(* Logix 5000 project; controller _GigaDiscovery vendor 1 type 14 code 244 rev 35.11; software revision 35.03; part 4 of 23 *)
(* tags used below, declared in another part *)
   Clock : DINT;   // Base tempi 10 milli sec
   Current_TimeInStation : DINT;
   Cycle_End_Timer : TIMER;
   Cycle_Timing : TIMER;
   Gates_Open_Permissive : Permissive;
   HMI_Angle : REAL;
   HMI_button_addtoindex : BOOL;
   HMI_button_subtracttoindex : BOOL;
   HMI_Current_Screen : DINT;
   HMI_Disable_external_acces : BOOL;   // ROUTER A72A07D Disable external acces
   HMI_Enable_external_acces : BOOL;   // ROUTER A72A07D Eneble external acces
   HMI_JM_Stats_Hist : Run_Count_Hist_JM[10];
   HMI_Lamp_Test : BOOL;
   HMI_Remote_Display : DINT;   // Display control 0 = operator 0 <> PLC
   HMI_Remote_Status : DINT;   // 0 = Disabled 1 = Enable but not remote control 2 = Remote control active
   HMI_Update_Time : BOOL;
   I_Light_Selector : BOOL;   // Light Selector Switch -S30408F
   I_OCC_Operator_Enable_Key : BOOL;   // OCC Console Enabled -S30305F
   I_Remote_Connection_Enabled : BOOL;   // Remote Connection active ROUTER eWON K74A04E
   index_for_stats_hist : DINT;
   Life_of_Machine : Life_of_Machine;
   No_Sfty : Std_to_Sfty;
   O_Enable_Remote_Connection : BOOL;   // ROUTER A72A07D Eneble external acces
   O_Front_Leg_Light : BOOL;   // Fron leg and front light signal -K3204H
   O_Gondola_Pendolum_Light : BOOL;   // Gondola and pendulum light signal -K3206H
   O_Rear_Leg_Light : BOOL;   // Rear leg and rear light signal -K3202H
   Platform_Close_Cycle : Sequencer;
   Platform_Close_Permissive : Permissive;
   Platform_Open_Cycle : Sequencer;
   Platform_Open_Permissive : Permissive;
   PltaformClosed_CycleComplete : BOOL;   // Piattaforme chiuse e ciclo completato
   PltaformOpeneded_CycleComplete : BOOL;   // Rilevazione Piattaforme aperte con ciclo Completato
   Previous_TimeInStation : DINT;
   ProofTest_Req : BOOL;
   RESTRAINTS_Closed : BOOL;   // All RESTRAINTS Closed
   RESTRAINTS_Closing : BOOL;
   Restraints_Cycle : Sequencer;
   RESTRAINTS_Opening : BOOL;
   Restraints_Permissive : Permissive;
   Restraints_Permissive_Ok : BOOL;
   Start_Permissive : Permissive;
   Start_Stop_Cycle : Sequencer;
   Start_TOF : TIMER;
   Stats_Times : DINT[30];
   TimeInStation_Count_Daily : COUNTER;
   TimeInStation_Count_Hourly : COUNTER;
   TimeInStation_Timer : TIMER;   // 10 min 600 sec
   Timers : TIMER[32];
   To_Sfty : Std_to_Sfty;

        [68].time_avg[17] := 29, [68].time_avg[18] := 26, [69].date[0] := -2, [69].date[1] := 1, [69].date[2] := 11, [69].runs[0] := 114, [69].runs[7] := 7, [69].runs[9] := 2, [69].runs[10] := 8, [69].runs[11] := 3, [69].runs[13] := 6, [69].runs[14] := 11, [69].time_avg[0] := 84, [69].time_avg[2] := 22683, [69].time_avg[4] := 28480, [69].time_avg[5] := 22361, [69].time_avg[7] := 107, [69].time_avg[11] := 24, [69].time_avg[13] := 70, [69].time_avg[14] := 104, [70].date[0] := -2, [70].date[1] := 1, [70].date[2] := 8, [70].runs[0] := 19, [70].runs[23] := 3, [70].time_avg[0] := 35, [70].time_avg[4] := 23240, [70].time_avg[5] := 22361, [71].date[0] := -2, [71].date[1] := 1, [71].date[2] := 7, [71].runs[0] := 30, [71].runs[20] := 2, [71].runs[21] := 6, [71].runs[22] := 1, [71].time_avg[0] := 199, [71].time_avg[4] := 23240, [71].time_avg[5] := 22361, [71].time_avg[21] := 199, [72].date[0] := -2, [72].date[1] := 1, [72].date[2] := 6, [72].runs[0] := 30, [72].time_avg[4] := 23240, [72].time_avg[5] := 22361, [73].date[0] := -2, [73].date[1] := 1, [73].date[2] := 5, [73].runs[0] := 4, [73].runs[23] := 1, [73].time_avg[4] := 23240, [73].time_avg[5] := 22361, [74].date[0] := 19, [74].date[1] := 9, [74].date[2] := 3, [74].runs[0] := 62, [74].runs[7] := 1, [74].runs[9] := 3, [74].runs[10] := 4, [74].runs[11] := 7,
        [74].runs[12] := 7, [74].runs[13] := 9, [74].runs[14] := 7, [74].runs[15] := 8, [74].runs[16] := 7, [74].runs[17] := 8, [74].runs[18] := 1, [74].runs[21] := 1, [74].time_avg[0] := 211, [74].time_avg[2] := 5236, [74].time_avg[3] := 12461, [74].time_avg[4] := 23240, [74].time_avg[5] := 22361, [74].time_avg[12] := 175, [74].time_avg[13] := 206, [74].time_avg[17] := 252, [74].time_avg[18] := 206, [74].time_avg[21] := 206, [75].date[0] := 19, [75].date[1] := 9, [75].date[2] := 2, [75].runs[0] := 70, [75].runs[7] := 1, [75].runs[9] := 4, [75].runs[10] := 3, [75].runs[12] := 6, [75].runs[13] := 7, [75].runs[14] := 5, [75].runs[15] := 9, [75].runs[16] := 7, [75].runs[17] := 2, [75].runs[18] := 8, [75].runs[19] := 9, [75].runs[20] := 8, [75].runs[21] := 1, [75].time_avg[0] := 186, [75].time_avg[2] := 5622, [75].time_avg[3] := 14544, [75].time_avg[4] := 20279, [75].time_avg[5] := 21563, [75].time_avg[10] := 214, [75].time_avg[12] := 152, [75].time_avg[13] := 173, [75].time_avg[14] := 183, [75].time_avg[15] := 191, [75].time_avg[16] := 193, [75].time_avg[17] := 150, [75].time_avg[18] := 177, [75].time_avg[19] := 190, [75].time_avg[20] := 190, [75].time_avg[21] := 370, [76].date[0] := 19, [76].date[1] := 9, [76].date[2] := 1, [76].runs[0] := 118, [76].runs[7] := 1, [76].runs[8] := 4, [76].runs[9] := 9, [76].runs[10] := 8, [76].runs[11] := 8,
        [76].runs[12] := 7, [76].runs[13] := 5, [76].runs[14] := 8, [76].runs[15] := 8, [76].runs[16] := 9, [76].runs[17] := 8, [76].runs[18] := 8, [76].runs[19] := 8, [76].runs[20] := 11, [76].runs[21] := 9, [76].runs[22] := 7, [76].time_avg[0] := 197, [76].time_avg[2] := 7812, [76].time_avg[3] := 8907, [76].time_avg[4] := 17438, [76].time_avg[5] := 20839, [76].time_avg[11] := 228, [76].time_avg[12] := 233, [76].time_avg[15] := 183, [76].time_avg[16] := 195, [76].time_avg[17] := 218, [76].time_avg[18] := 219, [76].time_avg[19] := 279, [76].time_avg[20] := 132, [76].time_avg[21] := 181, [76].time_avg[22] := 154, [77].date[0] := 19, [77].date[1] := 8, [77].date[2] := 31, [77].runs[0] := 121, [77].runs[7] := 1, [77].runs[9] := 6, [77].runs[10] := 11, [77].runs[11] := 8, [77].runs[12] := 9, [77].runs[13] := 9, [77].runs[14] := 9, [77].runs[15] := 8, [77].runs[16] := 9, [77].runs[17] := 9, [77].runs[18] := 9, [77].runs[19] := 9, [77].runs[20] := 10, [77].runs[21] := 8, [77].runs[22] := 6, [77].time_avg[0] := 193, [77].time_avg[2] := 4893, [77].time_avg[3] := 10185, [77].time_avg[4] := 20961, [77].time_avg[5] := 18600, [77].time_avg[10] := 199, [77].time_avg[11] := 202, [77].time_avg[12] := 189, [77].time_avg[13] := 205, [77].time_avg[14] := 168, [77].time_avg[15] := 213, [77].time_avg[16] := 188, [77].time_avg[17] := 210, [77].time_avg[18] := 201, [77].time_avg[19] := 185,
        [77].time_avg[20] := 174, [77].time_avg[21] := 198, [77].time_avg[22] := 164, [78].date[0] := 19, [78].date[1] := 8, [78].date[2] := 30, [78].runs[0] := 102, [78].runs[7] := 1, [78].runs[9] := 4, [78].runs[10] := 4, [78].runs[11] := 8, [78].runs[12] := 9, [78].runs[13] := 8, [78].runs[14] := 8, [78].runs[15] := 9, [78].runs[16] := 8, [78].runs[17] := 7, [78].runs[18] := 6, [78].runs[19] := 9, [78].runs[20] := 9, [78].runs[21] := 8, [78].runs[22] := 4, [78].time_avg[0] := 212, [78].time_avg[2] := 6981, [78].time_avg[3] := 13438, [78].time_avg[4] := 22920, [78].time_avg[5] := 22402, [78].time_avg[11] := 206, [78].time_avg[12] := 233, [78].time_avg[13] := 225, [78].time_avg[14] := 202, [78].time_avg[15] := 222, [78].time_avg[16] := 214, [78].time_avg[17] := 168, [78].time_avg[18] := 226, [78].time_avg[19] := 184, [78].time_avg[20] := 240, [78].time_avg[21] := 205, [78].time_avg[22] := 200, [79].date[0] := 19, [79].date[1] := 8, [79].date[2] := 29, [79].runs[0] := 108, [79].runs[9] := 4, [79].runs[10] := 5, [79].runs[11] := 9, [79].runs[12] := 10, [79].runs[13] := 10, [79].runs[14] := 10, [79].runs[15] := 8, [79].runs[16] := 9, [79].runs[17] := 10, [79].runs[18] := 9, [79].runs[19] := 9, [79].runs[20] := 9, [79].runs[21] := 5, [79].time_avg[0] := 182, [79].time_avg[2] := 4017, [79].time_avg[3] := 9797, [79].time_avg[4] := 23082,
        [79].time_avg[5] := 18998, [79].time_avg[10] := 174, [79].time_avg[11] := 200, [79].time_avg[12] := 157, [79].time_avg[13] := 156, [79].time_avg[14] := 151, [79].time_avg[15] := 216, [79].time_avg[16] := 184, [79].time_avg[17] := 179, [79].time_avg[18] := 206, [79].time_avg[19] := 187, [79].time_avg[20] := 186, [79].time_avg[21] := 214, [80].date[0] := 19, [80].date[1] := 8, [80].date[2] := 28, [80].runs[0] := 107, [80].runs[7] := 2, [80].runs[8] := 5, [80].runs[9] := 11, [80].runs[10] := 6, [80].runs[11] := 9, [80].runs[12] := 9, [80].runs[13] := 10, [80].runs[14] := 9, [80].runs[15] := 7, [80].runs[16] := 9, [80].runs[17] := 9, [80].runs[18] := 8, [80].runs[19] := 9, [80].runs[20] := 8, [80].runs[21] := 1, [80].time_avg[0] := 204, [80].time_avg[2] := 4432, [80].time_avg[3] := 11019, [80].time_avg[4] := 18000, [80].time_avg[5] := 22000, [80].time_avg[10] := 191, [80].time_avg[11] := 184, [80].time_avg[12] := 190, [80].time_avg[13] := 174, [80].time_avg[14] := 198, [80].time_avg[15] := 270, [80].time_avg[16] := 203, [80].time_avg[17] := 194, [80].time_avg[18] := 256, [80].time_avg[19] := 195, [80].time_avg[20] := 206, [80].time_avg[21] := 186, [81].date[0] := 19, [81].date[1] := 8, [81].date[2] := 27, [81].runs[0] := 114, [81].runs[7] := 1, [81].runs[9] := 4, [81].runs[10] := 5, [81].runs[11] := 9, [81].runs[12] := 8, [81].runs[13] := 8, [81].runs[14] := 9,
        [81].runs[15] := 11, [81].runs[16] := 10, [81].runs[17] := 11, [81].runs[18] := 11, [81].runs[19] := 12, [81].runs[20] := 9, [81].runs[21] := 6, [81].time_avg[0] := 146, [81].time_avg[2] := 5205, [81].time_avg[3] := 8324, [81].time_avg[4] := 51040, [81].time_avg[5] := 27563, [81].time_avg[10] := 152, [81].time_avg[11] := 179, [81].time_avg[12] := 150, [81].time_avg[13] := 187, [81].time_avg[14] := 179, [81].time_avg[15] := 142, [81].time_avg[16] := 146, [81].time_avg[17] := 112, [81].time_avg[18] := 141, [81].time_avg[19] := 93, [81].time_avg[20] := 163, [81].time_avg[21] := 149, [82].date[0] := 19, [82].date[1] := 8, [82].date[2] := 26, [82].runs[0] := 110, [82].runs[7] := 1, [82].runs[9] := 4, [82].runs[10] := 5, [82].runs[11] := 8, [82].runs[12] := 9, [82].runs[13] := 10, [82].runs[14] := 10, [82].runs[15] := 9, [82].runs[16] := 10, [82].runs[17] := 10, [82].runs[18] := 9, [82].runs[19] := 10, [82].runs[20] := 10, [82].runs[21] := 5, [82].time_avg[0] := 168, [82].time_avg[2] := 4284, [82].time_avg[3] := 14914, [82].time_avg[4] := 18760, [82].time_avg[5] := 19159, [82].time_avg[10] := 159, [82].time_avg[11] := 212, [82].time_avg[12] := 159, [82].time_avg[13] := 168, [82].time_avg[14] := 162, [82].time_avg[15] := 181, [82].time_avg[16] := 170, [82].time_avg[17] := 150, [82].time_avg[18] := 164, [82].time_avg[19] := 159, [82].time_avg[20] := 161, [82].time_avg[21] := 183, [83].date[0] := 19,
        [83].date[1] := 8, [83].date[2] := 25, [83].runs[0] := 116, [83].runs[7] := 1, [83].runs[9] := 4, [83].runs[10] := 4, [83].runs[11] := 9, [83].runs[12] := 9, [83].runs[13] := 9, [83].runs[14] := 11, [83].runs[15] := 10, [83].runs[16] := 9, [83].runs[17] := 9, [83].runs[18] := 7, [83].runs[19] := 11, [83].runs[20] := 9, [83].runs[21] := 10, [83].runs[22] := 4, [83].time_avg[0] := 171, [83].time_avg[2] := 3326, [83].time_avg[3] := 10694, [83].time_avg[4] := 30960, [83].time_avg[5] := 24322, [83].time_avg[10] := 258, [83].time_avg[11] := 206, [83].time_avg[12] := 166, [83].time_avg[13] := 166, [83].time_avg[14] := 133, [83].time_avg[15] := 149, [83].time_avg[16] := 187, [83].time_avg[17] := 204, [83].time_avg[18] := 204, [83].time_avg[19] := 143, [83].time_avg[20] := 164, [83].time_avg[21] := 145, [83].time_avg[22] := 212, [84].date[0] := 19, [84].date[1] := 8, [84].date[2] := 24, [84].runs[0] := 116, [84].runs[7] := 1, [84].runs[9] := 4, [84].runs[10] := 5, [84].runs[11] := 9, [84].runs[12] := 9, [84].runs[13] := 9, [84].runs[14] := 9, [84].runs[15] := 10, [84].runs[16] := 9, [84].runs[17] := 10, [84].runs[18] := 9, [84].runs[19] := 10, [84].runs[20] := 9, [84].runs[21] := 8, [84].runs[22] := 5, [84].time_avg[0] := 173, [84].time_avg[2] := 6434, [84].time_avg[3] := 9546, [84].time_avg[4] := 19840, [84].time_avg[5] := 19601,
        [84].time_avg[10] := 183, [84].time_avg[11] := 176, [84].time_avg[12] := 189, [84].time_avg[13] := 198, [84].time_avg[14] := 193, [84].time_avg[15] := 154, [84].time_avg[16] := 205, [84].time_avg[17] := 165, [84].time_avg[18] := 168, [84].time_avg[19] := 167, [84].time_avg[20] := 143, [84].time_avg[21] := 164, [84].time_avg[22] := 139, [85].date[0] := 19, [85].date[1] := 8, [85].date[2] := 23, [85].runs[0] := 108, [85].runs[7] := 1, [85].runs[9] := 4, [85].runs[10] := 3, [85].runs[11] := 10, [85].runs[12] := 9, [85].runs[13] := 8, [85].runs[14] := 9, [85].runs[15] := 10, [85].runs[16] := 9, [85].runs[17] := 9, [85].runs[18] := 8, [85].runs[19] := 9, [85].runs[20] := 9, [85].runs[21] := 8, [85].runs[22] := 2, [85].time_avg[0] := 204, [85].time_avg[2] := 6887, [85].time_avg[3] := 14477, [85].time_avg[4] := 20521, [85].time_avg[5] := 36240, [85].time_avg[10] := 221, [85].time_avg[11] := 190, [85].time_avg[12] := 186, [85].time_avg[13] := 191, [85].time_avg[14] := 226, [85].time_avg[15] := 161, [85].time_avg[16] := 185, [85].time_avg[17] := 211, [85].time_avg[18] := 232, [85].time_avg[19] := 218, [85].time_avg[20] := 196, [85].time_avg[21] := 251, [85].time_avg[22] := 235, [86].date[0] := 19, [86].date[1] := 8, [86].date[2] := 22, [86].runs[0] := 108, [86].runs[9] := 4, [86].runs[10] := 5, [86].runs[11] := 10, [86].runs[12] := 9, [86].runs[13] := 11, [86].runs[14] := 9,
        [86].runs[15] := 10, [86].runs[16] := 9, [86].runs[17] := 10, [86].runs[18] := 8, [86].runs[19] := 10, [86].runs[20] := 9, [86].runs[21] := 3, [86].time_avg[0] := 162, [86].time_avg[2] := 5022, [86].time_avg[3] := 11042, [86].time_avg[4] := 16840, [86].time_avg[5] := 22478, [86].time_avg[10] := 152, [86].time_avg[11] := 173, [86].time_avg[12] := 166, [86].time_avg[13] := 153, [86].time_avg[14] := 137, [86].time_avg[15] := 192, [86].time_avg[16] := 160, [86].time_avg[17] := 147, [86].time_avg[18] := 177, [86].time_avg[19] := 145, [86].time_avg[20] := 166, [86].time_avg[21] := 190, [87].date[0] := 19, [87].date[1] := 8, [87].date[2] := 21, [87].runs[0] := 110, [87].runs[9] := 5, [87].runs[10] := 5, [87].runs[11] := 9, [87].runs[12] := 8, [87].runs[13] := 10, [87].runs[14] := 10, [87].runs[15] := 10, [87].runs[16] := 10, [87].runs[17] := 9, [87].runs[18] := 10, [87].runs[19] := 8, [87].runs[20] := 9, [87].runs[21] := 6, [87].time_avg[0] := 174, [87].time_avg[2] := 5028, [87].time_avg[3] := 12622, [87].time_avg[4] := 18641, [87].time_avg[5] := 20757, [87].time_avg[9] := 267, [87].time_avg[10] := 158, [87].time_avg[11] := 186, [87].time_avg[12] := 162, [87].time_avg[13] := 179, [87].time_avg[14] := 156, [87].time_avg[15] := 147, [87].time_avg[16] := 154, [87].time_avg[17] := 158, [87].time_avg[18] := 185, [87].time_avg[19] := 180, [87].time_avg[20] := 236, [87].time_avg[21] := 167, [88].date[0] := 19,
        [88].date[1] := 8, [88].date[2] := 19, [88].runs[0] := 172, [88].runs[7] := 1, [88].runs[9] := 1, [88].runs[10] := 7, [88].runs[11] := 9, [88].runs[12] := 10, [88].runs[13] := 10, [88].runs[14] := 10, [88].runs[15] := 10, [88].runs[16] := 9, [88].runs[17] := 9, [88].runs[18] := 10, [88].runs[19] := 11, [88].runs[20] := 10, [88].runs[21] := 8, [88].time_avg[0] := 159, [88].time_avg[2] := 5010, [88].time_avg[3] := 9465, [88].time_avg[4] := 20080, [88].time_avg[5] := 17563, [88].time_avg[10] := 264, [88].time_avg[11] := 192, [88].time_avg[12] := 158, [88].time_avg[13] := 167, [88].time_avg[14] := 165, [88].time_avg[15] := 148, [88].time_avg[16] := 206, [88].time_avg[17] := 174, [88].time_avg[18] := 142, [88].time_avg[19] := 133, [88].time_avg[20] := 165, [88].time_avg[21] := 129, [89].date[0] := 19, [89].date[1] := 8, [89].date[2] := 18, [89].runs[0] := 116, [89].runs[7] := 1, [89].runs[10] := 8, [89].runs[11] := 10, [89].runs[12] := 10, [89].runs[13] := 9, [89].runs[14] := 10, [89].runs[15] := 11, [89].runs[16] := 4, [89].runs[17] := 9, [89].runs[18] := 10, [89].runs[19] := 10, [89].runs[20] := 9, [89].runs[21] := 11, [89].runs[22] := 4, [89].time_avg[0] := 160, [89].time_avg[2] := 4655, [89].time_avg[3] := 12877, [89].time_avg[4] := 21363, [89].time_avg[5] := 26439, [89].time_avg[10] := 166, [89].time_avg[11] := 166, [89].time_avg[12] := 161,
        [89].time_avg[13] := 187, [89].time_avg[14] := 165, [89].time_avg[15] := 133, [89].time_avg[16] := 160, [89].time_avg[17] := 161, [89].time_avg[18] := 173, [89].time_avg[19] := 149, [89].time_avg[20] := 175, [89].time_avg[21] := 139, [89].time_avg[22] := 162, [90].date[0] := 19, [90].date[1] := 8, [90].date[2] := 17, [90].runs[0] := 129, [90].runs[7] := 1, [90].runs[9] := 4, [90].runs[10] := 4, [90].runs[11] := 10, [90].runs[12] := 9, [90].runs[13] := 10, [90].runs[14] := 10, [90].runs[15] := 9, [90].runs[16] := 10, [90].runs[17] := 10, [90].runs[18] := 7, [90].runs[19] := 9, [90].runs[20] := 8, [90].runs[21] := 9, [90].runs[22] := 10, [90].runs[23] := 8, [90].time_avg[0] := 182, [90].time_avg[2] := 4196, [90].time_avg[3] := 11369, [90].time_avg[4] := 22122, [90].time_avg[5] := 21841, [90].time_avg[10] := 197, [90].time_avg[11] := 174, [90].time_avg[12] := 191, [90].time_avg[13] := 174, [90].time_avg[14] := 150, [90].time_avg[15] := 171, [90].time_avg[16] := 159, [90].time_avg[17] := 162, [90].time_avg[18] := 179, [90].time_avg[19] := 213, [90].time_avg[20] := 216, [90].time_avg[21] := 192, [90].time_avg[22] := 182, [90].time_avg[23] := 211, [91].date[0] := 19, [91].date[1] := 8, [91].date[2] := 16, [91].runs[0] := 110, [91].runs[7] := 1, [91].runs[9] := 4, [91].runs[10] := 6, [91].runs[11] := 10, [91].runs[12] := 8, [91].runs[13] := 9, [91].runs[14] := 3,
        [91].runs[15] := 10, [91].runs[16] := 10, [91].runs[17] := 10, [91].runs[18] := 9, [91].runs[19] := 9, [91].runs[20] := 9, [91].runs[21] := 10, [91].runs[22] := 2, [91].time_avg[0] := 167, [91].time_avg[2] := 5926, [91].time_avg[3] := 9632, [91].time_avg[4] := 23480, [91].time_avg[5] := 18838, [91].time_avg[10] := 161, [91].time_avg[11] := 149, [91].time_avg[12] := 156, [91].time_avg[13] := 170, [91].time_avg[15] := 151, [91].time_avg[16] := 156, [91].time_avg[17] := 158, [91].time_avg[18] := 203, [91].time_avg[19] := 192, [91].time_avg[20] := 185, [91].time_avg[21] := 150, [91].time_avg[22] := 195, [92].date[0] := 19, [92].date[1] := 8, [92].date[2] := 15, [92].runs[0] := 113, [92].runs[7] := 1, [92].runs[9] := 4, [92].runs[10] := 5, [92].runs[11] := 9, [92].runs[12] := 9, [92].runs[13] := 9, [92].runs[14] := 9, [92].runs[15] := 10, [92].runs[16] := 10, [92].runs[17] := 9, [92].runs[18] := 10, [92].runs[19] := 9, [92].runs[20] := 10, [92].runs[21] := 9, [92].time_avg[0] := 174, [92].time_avg[2] := 4980, [92].time_avg[3] := 11102, [92].time_avg[4] := 19122, [92].time_avg[5] := 22677, [92].time_avg[10] := 180, [92].time_avg[11] := 184, [92].time_avg[12] := 201, [92].time_avg[13] := 188, [92].time_avg[14] := 179, [92].time_avg[15] := 164, [92].time_avg[16] := 165, [92].time_avg[17] := 189, [92].time_avg[18] := 169, [92].time_avg[19] := 168, [92].time_avg[20] := 159, [92].time_avg[21] := 153,
        [93].date[0] := 19, [93].date[1] := 8, [93].date[2] := 14, [93].runs[0] := 110, [93].runs[7] := 1, [93].runs[9] := 4, [93].runs[10] := 5, [93].runs[11] := 9, [93].runs[12] := 10, [93].runs[13] := 10, [93].runs[14] := 10, [93].runs[15] := 10, [93].runs[16] := 10, [93].runs[17] := 8, [93].runs[18] := 10, [93].runs[19] := 10, [93].runs[20] := 8, [93].runs[21] := 5, [93].time_avg[0] := 170, [93].time_avg[2] := 3396, [93].time_avg[3] := 11574, [93].time_avg[4] := 19402, [93].time_avg[5] := 24403, [93].time_avg[10] := 164, [93].time_avg[11] := 183, [93].time_avg[12] := 161, [93].time_avg[13] := 163, [93].time_avg[14] := 151, [93].time_avg[15] := 150, [93].time_avg[16] := 168, [93].time_avg[17] := 227, [93].time_avg[18] := 179, [93].time_avg[19] := 161, [93].time_avg[20] := 173, [93].time_avg[21] := 178, [94].date[0] := 19, [94].date[1] := 8, [94].date[2] := 13, [94].runs[0] := 99, [94].runs[7] := 1, [94].runs[9] := 4, [94].runs[10] := 4, [94].runs[11] := 11, [94].runs[12] := 8, [94].runs[13] := 5, [94].runs[14] := 9, [94].runs[15] := 8, [94].runs[16] := 10, [94].runs[17] := 9, [94].runs[18] := 8, [94].runs[19] := 9, [94].runs[20] := 8, [94].runs[21] := 5, [94].time_avg[0] := 185, [94].time_avg[2] := 4905, [94].time_avg[3] := 9992, [94].time_avg[4] := 19077, [94].time_avg[5] := 20762, [94].time_avg[10] := 183, [94].time_avg[11] := 135,
        [94].time_avg[12] := 171, [94].time_avg[13] := 195, [94].time_avg[14] := 209, [94].time_avg[15] := 185, [94].time_avg[16] := 185, [94].time_avg[17] := 186, [94].time_avg[18] := 200, [94].time_avg[19] := 175, [94].time_avg[20] := 224, [94].time_avg[21] := 204, [95].date[0] := 19, [95].date[1] := 8, [95].date[2] := 12, [95].runs[0] := 118, [95].runs[8] := 1, [95].runs[9] := 6, [95].runs[10] := 5, [95].runs[11] := 10, [95].runs[12] := 11, [95].runs[13] := 10, [95].runs[14] := 8, [95].runs[15] := 10, [95].runs[16] := 10, [95].runs[17] := 10, [95].runs[18] := 10, [95].runs[19] := 8, [95].runs[20] := 9, [95].runs[21] := 10, [95].time_avg[0] := 156, [95].time_avg[2] := 6366, [95].time_avg[3] := 11660, [95].time_avg[4] := 23243, [95].time_avg[5] := 28239, [95].time_avg[10] := 194, [95].time_avg[11] := 153, [95].time_avg[12] := 133, [95].time_avg[13] := 156, [95].time_avg[14] := 137, [95].time_avg[15] := 150, [95].time_avg[16] := 151, [95].time_avg[17] := 145, [95].time_avg[18] := 164, [95].time_avg[19] := 182, [95].time_avg[20] := 195, [95].time_avg[21] := 148, [96].date[0] := 19, [96].date[1] := 8, [96].date[2] := 11, [96].runs[0] := 123, [96].runs[7] := 1, [96].runs[9] := 4, [96].runs[10] := 8, [96].runs[11] := 10, [96].runs[12] := 11, [96].runs[13] := 10, [96].runs[14] := 7, [96].runs[15] := 11, [96].runs[16] := 9, [96].runs[17] := 10, [96].runs[18] := 9,
        [96].runs[19] := 11, [96].runs[20] := 8, [96].runs[21] := 9, [96].runs[22] := 5, [96].time_avg[0] := 157, [96].time_avg[2] := 4752, [96].time_avg[3] := 9692, [96].time_avg[4] := 19361, [96].time_avg[5] := 22281, [96].time_avg[10] := 173, [96].time_avg[11] := 141, [96].time_avg[12] := 142, [96].time_avg[13] := 141, [96].time_avg[14] := 179, [96].time_avg[15] := 138, [96].time_avg[16] := 183, [96].time_avg[17] := 147, [96].time_avg[18] := 191, [96].time_avg[19] := 146, [96].time_avg[20] := 167, [96].time_avg[21] := 162, [96].time_avg[22] := 167, [97].date[0] := 19, [97].date[1] := 8, [97].date[2] := 10, [97].runs[0] := 120, [97].runs[7] := 1, [97].runs[9] := 5, [97].runs[10] := 4, [97].runs[11] := 6, [97].runs[12] := 8, [97].runs[13] := 11, [97].runs[14] := 8, [97].runs[15] := 11, [97].runs[16] := 9, [97].runs[17] := 10, [97].runs[18] := 11, [97].runs[19] := 10, [97].runs[20] := 11, [97].runs[21] := 10, [97].runs[22] := 5, [97].time_avg[0] := 142, [97].time_avg[2] := 4697, [97].time_avg[3] := 8479, [97].time_avg[4] := 21362, [97].time_avg[5] := 36560, [97].time_avg[10] := 200, [97].time_avg[11] := 178, [97].time_avg[12] := 152, [97].time_avg[13] := 141, [97].time_avg[14] := 131, [97].time_avg[15] := 153, [97].time_avg[16] := 133, [97].time_avg[17] := 145, [97].time_avg[18] := 140, [97].time_avg[19] := 135, [97].time_avg[20] := 138, [97].time_avg[21] := 126, [97].time_avg[22] := 121, [98].date[0] := 19,
        [98].date[1] := 8, [98].date[2] := 9, [98].runs[0] := 119, [98].runs[7] := 1, [98].runs[9] := 5, [98].runs[10] := 5, [98].runs[11] := 8, [98].runs[12] := 9, [98].runs[13] := 8, [98].runs[14] := 11, [98].runs[15] := 11, [98].runs[16] := 8, [98].runs[17] := 10, [98].runs[18] := 9, [98].runs[19] := 11, [98].runs[20] := 9, [98].runs[21] := 10, [98].runs[22] := 4, [98].time_avg[0] := 151, [98].time_avg[2] := 4804, [98].time_avg[3] := 10881, [98].time_avg[4] := 800, [98].time_avg[5] := 21920, [98].time_avg[9] := 35, [98].time_avg[10] := 126, [98].time_avg[11] := 166, [98].time_avg[12] := 159, [98].time_avg[13] := 165, [98].time_avg[14] := 138, [98].time_avg[15] := 126, [98].time_avg[16] := 148, [98].time_avg[17] := 148, [98].time_avg[18] := 187, [98].time_avg[19] := 138, [98].time_avg[20] := 165, [98].time_avg[21] := 145, [98].time_avg[22] := 168, [99].date[0] := 19, [99].date[1] := 8, [99].date[2] := 8, [99].runs[0] := 93, [99].runs[7] := 1, [99].runs[9] := 4, [99].runs[10] := 4, [99].runs[11] := 9, [99].runs[12] := 9, [99].runs[13] := 9, [99].runs[14] := 8, [99].runs[15] := 9, [99].runs[16] := 9, [99].runs[17] := 2, [99].runs[18] := 5, [99].runs[19] := 8, [99].runs[20] := 9, [99].runs[21] := 7, [99].time_avg[0] := 156, [99].time_avg[2] := 5998, [99].time_avg[3] := 7111, [99].time_avg[4] := 17880, [99].time_avg[5] := 21321,
        [99].time_avg[10] := 153, [99].time_avg[11] := 154, [99].time_avg[12] := 146, [99].time_avg[13] := 139, [99].time_avg[14] := 173, [99].time_avg[15] := 152, [99].time_avg[16] := 160, [99].time_avg[17] := 133, [99].time_avg[18] := 182, [99].time_avg[19] := 147, [99].time_avg[20] := 148, [99].time_avg[21] := 188);
   MINUTE : DINT := 40;   // Minute
   MONTH : DINT := 12;   // Month
   MUL_01 : FBD_MATH := (SourceB := 1.13);
   Opening_CyclePlatTimes : DINT[20] := ([1] := 22393, [2] := 3119, [3] := 6800, [4] := 18122, [5] := 19079, [6] := 22361, [9] := 11322, [10] := 11039);
        [14]   // daily overall avg
        [13]   // daily overall total
   Os : DINT := 1280;
   Runs_DAILY : DINT := 11;   // Daily Total
   Runs_HOURLY : DINT := 3;   // Hourly Total
   Runs_LAST_YEARLY : DINT := 352;   // Last Year Total
   Runs_YEARLY : DINT := 1755;   // Yearly Total
   SECOND : DINT := 55;   // Second
   STATS_ONS : DINT := 24;
        .5   // ONS Stats 5 New Hour
        .4   // ONS Stats 4 New Day
        .10   // ONS Stats 10 Run Time
        .21   // ONS Stats 21
        .22   // ONS Stats 22
        .23   // ONS Stats 23
        .24   // ONS Stats 24
        .11   // ONS Stats 11 Screen RuntCt
        .2   // ONS Stats 2 Increment Count
        .9   // ONS Stas 9 End TImeInStation
        .1   // ONS Stats 1 Count Dispatch
        .25   // ONS Stats 25
        .3   // ONS Stats 3 New Year
        .26   // ONS Stats 26
        .27   // ONS Stats 27
        .28   // ONS Stats 28
        .12   // ONS Stats 12 Add Index
        .29   // ONS Stats 29
        .8   // ONS Stats 8 Start TimeInStation
        .30   // ONS Stats 30
        .13   // ONS Stats 13 Sub Index
   STATS_Plat_ONS : DINT;
        .11   // ONS Stats 11 Before Cycle Platform Open Avail
        .3   // ONS Stats 3 End Cycle Platform Close Pushed
        .14   // ONS Stats 14 Before Cycle Platform All Good
        .1   // ONS Stats 1 End Cycle Platform Avail
        .4   // ONS Stats 4 End Cycle Platform All Good
        .5   // ONS Stats 5 End Cycle Lever Disabled
        .2   // ONS Stats 2 End Cycle Lever Enabled
        .15   // ONS Stats 15 Before Cycle Lever Disabled
        .16   // ONS Stats 15 Before Cycle Ride Started
        .12   // ONS Stats 12 Before Cycle Lever Enabled
        .13   // ONS Stats 13 Before Cycle Platform Open Pushed
        .6   // ONS Stats 6 Gates and Bars Open
   Time_Date : DINT[7] := ([0] := 2025, [1] := 12, [2] := 1, [3] := 19, [4] := 40, [5] := 55, [6] := 815141);
   Timer : TIMER[10] := ([0].PRE := 10000, [1].PRE := 10000, [1].ACC := 10000, [2].PRE := 2000, [3].PRE := 2000, [3].ACC := 2000, [3].EN := 1, [3].DN := 1, [4].PRE := 1000, [5].PRE := 600000, [5].EN := 1, [5].DN := 1, [6].PRE := 660000, [6].EN := 1, [6].DN := 1);
   Total_TimeInStation_Daily : DINT := 1244;
   Total_TimeInStation_Hourly : DINT := 606;
   Trigger : DINT;   // Triggers
        .5   // Trigger 5 Cycle Ended
        .2   // Trigger 2 Dispatch Start
        .20   // Trigger 20 Was Loading
        .1   // Trigger 1 TimeInStation Start
        .0   // Trigger 0 Dispatch Counted
   YEAR : DINT := 2025;   // Year
END_VAR

ROUTINE _01_Life_of_Machine   (* ladder *)
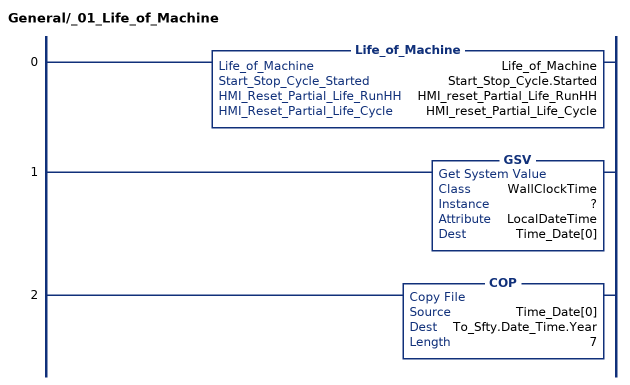
   [picture p37: General/_01_Life_of_Machine rungs 0-2]
   0: Life_of_Machine(Life_of_Machine,Start_Stop_Cycle.Started,HMI_reset_Partial_Life_RunHH,HMI_reset_Partial_Life_Cycle);
   1: GSV(WallClockTime,?,LocalDateTime,Time_Date[0]);
   2: COP(Time_Date[0],To_Sfty.Date_Time.Year,7);
END_ROUTINE

ROUTINE _02_Safety_Signature   (* ladder *)
END_ROUTINE

ROUTINE _03_Lights   (* ladder *)
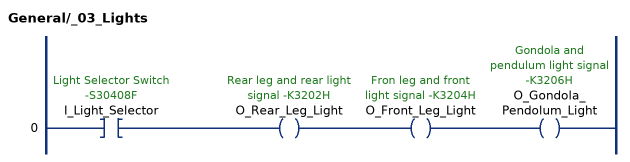
   0: XIC(I_Light_Selector)OTE(O_Rear_Leg_Light)OTE(O_Front_Leg_Light)OTE(O_Gondola_Pendolum_Light);
END_ROUTINE

ROUTINE _04_Router   (* ladder *)
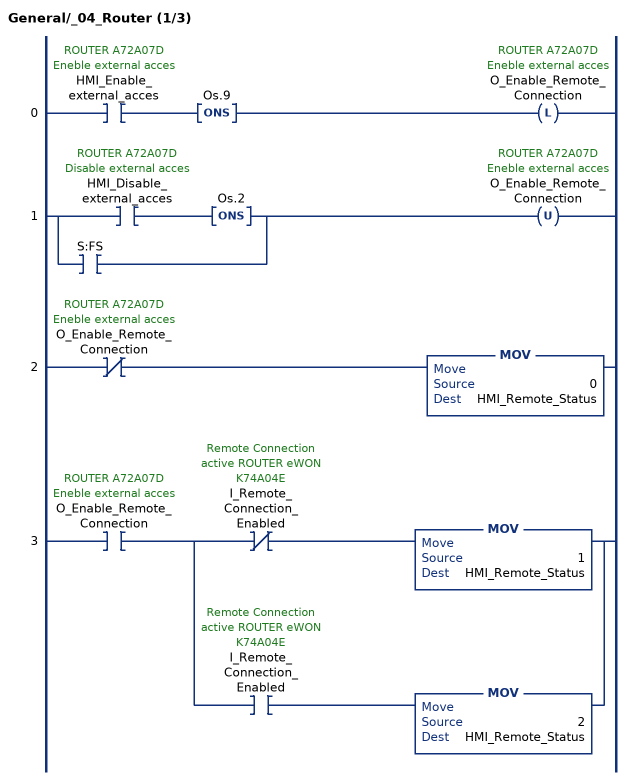
   0: XIC(HMI_Enable_external_acces)ONS(Os.9)OTL(O_Enable_Remote_Connection);
   1: [XIC(HMI_Disable_external_acces) ONS(Os.2) ,XIC(S:FS) ]OTU(O_Enable_Remote_Connection);
   2: XIO(O_Enable_Remote_Connection)MOV(0,HMI_Remote_Status);
   3: XIC(O_Enable_Remote_Connection)[XIO(I_Remote_Connection_Enabled) MOV(1,HMI_Remote_Status) ,XIC(I_Remote_Connection_Enabled) MOV(2,HMI_Remote_Status) ];
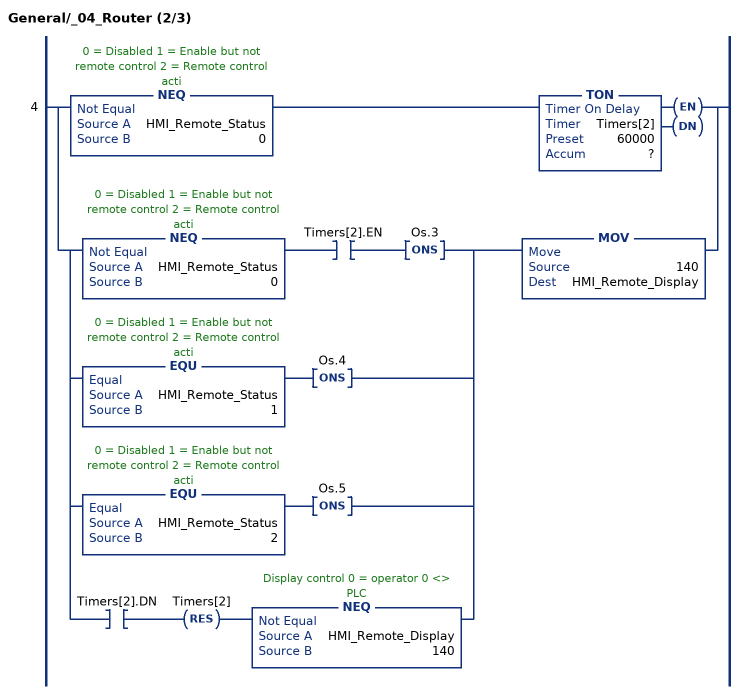
   4: [NEQ(HMI_Remote_Status,0) TON(Timers[2],?,?) ,[NEQ(HMI_Remote_Status,0) XIC(Timers[2].EN) ONS(Os.3) ,EQU(HMI_Remote_Status,1) ONS(Os.4) ,EQU(HMI_Remote_Status,2) ONS(Os.5) ,XIC(Timers[2].DN) RES(Timers[2]) NEQ(HMI_Remote_Display,140) ] MOV(140,HMI_Remote_Display) ];